
screen "MTA-CFGAvisosBAJA" 1280x800, template "Plantilla"
   TextField "Campo de texto_1" at 477,9 size 354x27; Text 'Configuración de avisos para Baja presión'
   TextField "Campo de texto_9" at 161,54 size 281x34; Text 'Avisos de BAJA PRESIÓN'
   IOField "Campo ES_1" at 295,105 size 130x30; Authorization "Administración de usuarios"; FormatPattern 999.99; Unit  bar
      ProcessValue <- "CFG-BajaHH"
   IOField "Campo ES_2" at 295,240 size 130x31; Authorization "Administración de usuarios"; FormatPattern 9999999; Unit  h
      ProcessValue <- "Varios_HorasMantMC061_1"
   IOField "Campo ES_3" at 295,195 size 130x31; Authorization "Administración de usuarios"; FormatPattern 9999999; Unit  h
      ProcessValue <- "Varios_HorasMantMC060_3"
   IOField "Campo ES_4" at 295,150 size 130x31; Authorization "Administración de usuarios"; FormatPattern 999.99; Unit  bar
      ProcessValue <- "CFG-BajaLL"
   IOField "Campo ES_5" at 295,285 size 130x30; Authorization "Administración de usuarios"; FormatPattern 9999999; Unit  h
      ProcessValue <- "Varios_HorasMantMC061_4"
   IOField "Campo ES_6" at 295,330 size 130x31; Authorization "Administración de usuarios"; FormatPattern 9999999; Unit  h
      ProcessValue <- "Varios_HorasMantMC062_2"
   IOField "Campo ES_7" at 295,375 size 130x31; Authorization "Administración de usuarios"; FormatPattern 9999999; Unit  h
      ProcessValue <- "Varios_HorasMantMC062_5"
   IOField "Campo ES_8" at 295,420 size 130x31; Authorization "Administración de usuarios"; FormatPattern 9999999; Unit  h
      ProcessValue <- "Varios_HorasMantMC063_3"
   TextField "Campo de texto_2" at 15,107 size 293x25; Text 'Presión Aviso límite de presión Máxima'
   TextField "Campo de texto_3" at 15,242 size 238x25; Text 'Tiempo Mant.#1 Comp. Sullair1'
   TextField "Campo de texto_6" at 15,197 size 248x25; Text 'Tiempo Mant. #3 Comp. Sullair2'
   TextField "Campo de texto_4" at 15,152 size 289x25; Text 'Presión Aviso límite de presión Mínima'
   TextField "Campo de texto_5" at 15,287 size 238x25; Text 'Tiempo Mant.#4 Comp. Sullair1'
   TextField "Campo de texto_7" at 15,332 size 238x25; Text 'Tiempo Mant.#2 Comp. Sullair0'
   TextField "Campo de texto_8" at 15,377 size 238x25; Text 'Tiempo Mant.#5 Comp. Sullair0'
   TextField "Campo de texto_10" at 15,422 size 231x25; Text 'Tiempo Mant.#3 Comp. Atlas3'
   IOField "Campo ES_9" at 295,465 size 130x30; Authorization "Administración de usuarios"; FormatPattern 9999999; Unit  h
      ProcessValue <- "Varios_HorasMantMC064_1"
   IOField "Campo ES_10" at 295,510 size 130x31; Authorization "Administración de usuarios"; FormatPattern 9999999; Unit  h
      ProcessValue <- "Varios_HorasMantMC064_4"
   IOField "Campo ES_11" at 295,555 size 130x31; Authorization "Administración de usuarios"; FormatPattern 9999999; Unit  h
      ProcessValue <- "Varios_HorasMantMS054_2"
   TextField "Campo de texto_11" at 15,467 size 231x25; Text 'Tiempo Mant.#1 Comp. Atlas2'
   TextField "Campo de texto_12" at 15,512 size 231x25; Text 'Tiempo Mant.#4 Comp. Atlas2'
   TextField "Campo de texto_13" at 15,557 size 232x25; Text 'Tiempo Mant. #2 Sec. Sullair 1'
   IOField "Campo ES_13" at 716,150 size 130x30; Authorization "Administración de usuarios"; FormatPattern 9999999; Unit  h
      ProcessValue <- "Varios_HorasMantMC060_1"
   IOField "Campo ES_14" at 716,105 size 130x31; Authorization "Administración de usuarios"; FormatPattern 999.99; Unit  bar
      ProcessValue <- "CFG-BajaH"
   IOField "Campo ES_15" at 716,195 size 130x31; Authorization "Administración de usuarios"; FormatPattern 9999999; Unit  h
      ProcessValue <- "Varios_HorasMantMC060_4"
   IOField "Campo ES_16" at 716,240 size 130x31; Authorization "Administración de usuarios"; FormatPattern 9999999; Unit  h
      ProcessValue <- "Varios_HorasMantMC061_2"
   IOField "Campo ES_17" at 716,285 size 130x30; Authorization "Administración de usuarios"; FormatPattern 9999999; Unit  h
      ProcessValue <- "Varios_HorasMantMC061_5"
   IOField "Campo ES_18" at 716,330 size 130x31; Authorization "Administración de usuarios"; FormatPattern 9999999; Unit  h
      ProcessValue <- "Varios_HorasMantMC062_3"
   IOField "Campo ES_19" at 716,375 size 130x31; Authorization "Administración de usuarios"; FormatPattern 9999999; Unit  h
      ProcessValue <- "Varios_HorasMantMC063_1"
   IOField "Campo ES_20" at 716,420 size 130x31; Authorization "Administración de usuarios"; FormatPattern 9999999; Unit  h
      ProcessValue <- "Varios_HorasMantMC063_4"
   TextField "Campo de texto_15" at 436,152 size 248x25; Text 'Tiempo Mant. #1 Comp. Sullair2'
   TextField "Campo de texto_16" at 436,107 size 247x25; Text 'Presión Aviso de presión elevada'
   TextField "Campo de texto_17" at 436,197 size 248x25; Text 'Tiempo Mant. #4 Comp. Sullair2'
   TextField "Campo de texto_18" at 436,242 size 238x25; Text 'Tiempo Mant.#2 Comp. Sullair1'
   TextField "Campo de texto_19" at 436,287 size 238x25; Text 'Tiempo Mant.#5 Comp. Sullair1'
   TextField "Campo de texto_20" at 436,332 size 238x25; Text 'Tiempo Mant.#3 Comp. Sullair0'
   TextField "Campo de texto_21" at 436,377 size 231x25; Text 'Tiempo Mant.#1 Comp. Atlas3'
   TextField "Campo de texto_22" at 436,422 size 231x25; Text 'Tiempo Mant.#4 Comp. Atlas3'
   IOField "Campo ES_21" at 716,465 size 130x30; Authorization "Administración de usuarios"; FormatPattern 9999999; Unit  h
      ProcessValue <- "Varios_HorasMantMC064_2"
   IOField "Campo ES_22" at 716,510 size 130x31; Authorization "Administración de usuarios"; FormatPattern 9999999; Unit  h
      ProcessValue <- "Varios_HorasMantMC064_5"
   IOField "Campo ES_23" at 716,555 size 130x31; Authorization "Administración de usuarios"; FormatPattern 9999999; Unit  h
      ProcessValue <- "Varios_UltimoMantMS055_1"
   TextField "Campo de texto_23" at 436,467 size 231x25; Text 'Tiempo Mant.#2 Comp. Atlas2'
   TextField "Campo de texto_24" at 436,512 size 231x25; Text 'Tiempo Mant.#5 Comp. Atlas2'
   TextField "Campo de texto_25" at 436,557 size 232x25; Text 'Tiempo Mant. #1 Sec. Sullair 2'
   IOField "Campo ES_25" at 1137,195 size 130x30; Authorization "Administración de usuarios"; FormatPattern 9999999; Unit  h
      ProcessValue <- "Varios_UltimoMantMC060_5"
   IOField "Campo ES_26" at 1137,150 size 130x31; Authorization "Administración de usuarios"; FormatPattern 9999999; Unit  h
      ProcessValue <- "Varios_HorasMantMC060_2"
   IOField "Campo ES_27" at 1137,105 size 130x31; Authorization "Administración de usuarios"; FormatPattern 999.99; Unit  bar
      ProcessValue <- "CFG-BajaL"
   IOField "Campo ES_28" at 1137,240 size 130x31; Authorization "Administración de usuarios"; FormatPattern 9999999; Unit  h
      ProcessValue <- "Varios_HorasMantMC061_3"
   IOField "Campo ES_29" at 1137,285 size 130x30; Authorization "Administración de usuarios"; FormatPattern 9999999; Unit  h
      ProcessValue <- "Varios_HorasMantMC062_1"
   IOField "Campo ES_30" at 1137,330 size 130x31; Authorization "Administración de usuarios"; FormatPattern 9999999; Unit  h
      ProcessValue <- "Varios_HorasMantMC062_4"
   IOField "Campo ES_31" at 1137,375 size 130x31; Authorization "Administración de usuarios"; FormatPattern 9999999; Unit  h
      ProcessValue <- "Varios_HorasMantMC063_2"
   IOField "Campo ES_32" at 1137,420 size 130x31; Authorization "Administración de usuarios"; FormatPattern 9999999; Unit  h
      ProcessValue <- "Varios_HorasMantMC063_5"
   TextField "Campo de texto_27" at 857,197 size 243x25; Text 'Tiempo Mant.#5 Comp. Sullair2'
   TextField "Campo de texto_28" at 857,152 size 248x25; Text 'Tiempo Mant. #2 Comp. Sullair2'
   TextField "Campo de texto_29" at 857,107 size 222x25; Text 'Presión Aviso de presión baja'
   TextField "Campo de texto_30" at 857,242 size 238x25; Text 'Tiempo Mant.#3 Comp. Sullair1'
   TextField "Campo de texto_31" at 857,287 size 238x25; Text 'Tiempo Mant.#1 Comp. Sullair0'
   TextField "Campo de texto_32" at 857,332 size 238x25; Text 'Tiempo Mant.#4 Comp. Sullair0'
   TextField "Campo de texto_33" at 857,377 size 231x25; Text 'Tiempo Mant.#2 Comp. Atlas3'
   TextField "Campo de texto_34" at 857,422 size 273x25; Text 'Tiempo mant. #5 compresor Atlas 3'
   IOField "Campo ES_33" at 1137,465 size 130x30; Authorization "Administración de usuarios"; FormatPattern 9999999; Unit  h
      ProcessValue <- "Varios_HorasMantMC064_3"
   IOField "Campo ES_34" at 1137,510 size 130x31; Authorization "Administración de usuarios"; FormatPattern 9999999; Unit  h
      ProcessValue <- "Varios_HorasMantMS054_1"
   IOField "Campo ES_35" at 1137,555 size 130x31; Authorization "Administración de usuarios"; FormatPattern 9999999; Unit  h
      ProcessValue <- "Varios_HorasMantMS055_2"
   TextField "Campo de texto_35" at 857,467 size 231x25; Text 'Tiempo Mant.#3 Comp. Atlas2'
   TextField "Campo de texto_36" at 857,512 size 232x25; Text 'Tiempo Mant. #1 Sec. Sullair 1'
   TextField "Campo de texto_37" at 857,557 size 232x25; Text 'Tiempo Mant. #2 Sec. Sullair 2'

screen "MTA-ChillersBombasEnvasado" 1280x800, template "Plantilla"
   TextField "Campo de texto_5" at 519,10 size 240x27; Text 'Chillers - Bombas Envasado'
   GraphicView "Visor de gráficos_3" at 944,375 size 64x103; Picture "Bomba"
   GraphicIOField "Plantilla_Campo ES gráfico_2" at 980,449 size 81x68; PictureList "Motor2"
      ProcessValue <- "AnimaciónMT009"
   SymbolicIOField "Campo ES simbólico_4" at 890,188 size 220x29; TextOff '0'; TextOn '1'; TextList "EstadoMotor"
      ProcessValue <- "AnimaciónMT009"
   TextField "Campo de texto_6" at 887,129 size 53x23; Text 'MT009'
   GraphicView "Visor de gráficos_4" at 702,375 size 64x103; Picture "Bomba"
   GraphicIOField "Plantilla_Campo ES gráfico_1" at 738,449 size 81x68; PictureList "Motor2"
      ProcessValue <- "AnimaciónMT010"
   SymbolicIOField "Campo ES simbólico_1" at 648,188 size 220x29; TextOff '0'; TextOn '1'; TextList "EstadoMotor"
      ProcessValue <- "AnimaciónMT010"
   TextField "Campo de texto_7" at 645,129 size 53x23; Text 'MT010'
   GraphicView "Visor de gráficos_6" at 216,375 size 64x103; Picture "Bomba"
   GraphicIOField "Plantilla_Campo ES gráfico_4" at 252,449 size 81x68; PictureList "Motor2"
      ProcessValue <- "AnimaciónMP013"
   SymbolicIOField "Campo ES simbólico_3" at 164,188 size 220x29; TextOff '0'; TextOn '1'; TextList "EstadoMotor"
      ProcessValue <- "AnimaciónMP013"
   TextField "Campo de texto_9" at 167,129 size 52x23; Text 'MP013'
   TextField "Campo de texto_19" at 645,160 size 195x18; Text 'Intercambiador Línea 1 y Manomec'
   GraphicView "Visor de gráficos_5" at 460,375 size 64x103; Picture "Bomba"
   GraphicIOField "Plantilla_Campo ES gráfico_3" at 496,449 size 81x68; PictureList "Motor2"
      ProcessValue <- "AnimaciónMP012"
   SymbolicIOField "Campo ES simbólico_2" at 406,188 size 220x29; TextOff '0'; TextOn '1'; TextList "EstadoMotor"
      ProcessValue <- "AnimaciónMP012"
   TextField "Campo de texto_8" at 403,129 size 52x23; Text 'MP012'
   TextField "Campo de texto_18" at 886,160 size 150x18; Text 'Intercambiador Línea 3 y 5'
   TextField "Campo de texto_16" at 407,161 size 150x18; Text 'Chillers Envasado - Principal'
   TextField "Campo de texto_17" at 165,161 size 146x18; Text 'Chillers Envasado - Backup'
   ScreenModuleView "ControlMotor-NoAUTO_1" at 916,230 size 171x108
      Guid_{11997190-67152} <- "DesMT009"
      Guid_{11997190-67156} <- "ParadaMT009"
      Guid_{11997190-67150} <- "HabMT009"
      Guid_{11997190-67154} <- "MarchaMT009"
   ScreenModuleView "ControlMotor-NoAUTO_2" at 676,230 size 171x108
      Guid_{11997190-67152} <- "DesMT010"
      Guid_{11997190-67156} <- "ParadaMT010"
      Guid_{11997190-67150} <- "HabMT010"
      Guid_{11997190-67154} <- "MarchaMT010"
   ScreenModuleView "ControlMotor-NoAUTO_3" at 431,230 size 171x108
      Guid_{11997190-67152} <- "DesMP012"
      Guid_{11997190-67156} <- "ParadaMP012"
      Guid_{11997190-67150} <- "HabMP012"
      Guid_{11997190-67154} <- "MarchaMP012"
   ScreenModuleView "ControlMotor-NoAUTO_4" at 191,230 size 171x108
      Guid_{11997190-67152} <- "DesMP013"
      Guid_{11997190-67156} <- "ParadaMP013"
      Guid_{11997190-67150} <- "HabMP013"
      Guid_{11997190-67154} <- "MarchaMP013"
   Button "Botón_1" at 1184,68 size 48x46; TextOff '?'
      on Click: ActivateScreen("MTA-AyudaMotores", 0)

screen "MTA-ChillersBombasSoplado" 1280x800, template "Plantilla"
   GraphicView "Visor de gráficos_3" at 944,375 size 64x103; Picture "Bomba"
   GraphicView "Visor de gráficos_4" at 702,375 size 64x103; Picture "Bomba"
   GraphicView "Visor de gráficos_6" at 216,375 size 64x103; Picture "Bomba"
   GraphicView "Visor de gráficos_5" at 460,375 size 64x103; Picture "Bomba"
   TextField "Campo de texto_5" at 530,10 size 221x27; Text 'Chillers - Bombas Soplado'
   GraphicIOField "Plantilla_Campo ES gráfico_2" at 980,449 size 81x68; PictureList "Motor2"
      ProcessValue <- "AnimaciónMT007"
   SymbolicIOField "Campo ES simbólico_4" at 890,188 size 220x29; TextOff '0'; TextOn '1'; TextList "EstadoMotor"
      ProcessValue <- "AnimaciónMT007"
   TextField "Campo de texto_6" at 887,129 size 53x23; Text 'MT007'
   GraphicIOField "Plantilla_Campo ES gráfico_1" at 738,449 size 81x68; PictureList "Motor2"
      ProcessValue <- "AnimaciónMT008"
   SymbolicIOField "Campo ES simbólico_1" at 648,188 size 220x29; TextOff '0'; TextOn '1'; TextList "EstadoMotor"
      ProcessValue <- "AnimaciónMT008"
   TextField "Campo de texto_7" at 645,129 size 53x23; Text 'MT008'
   GraphicIOField "Plantilla_Campo ES gráfico_4" at 252,449 size 81x68; PictureList "Motor2"
      ProcessValue <- "AnimaciónMP011"
   SymbolicIOField "Campo ES simbólico_3" at 164,188 size 220x29; TextOff '0'; TextOn '1'; TextList "EstadoMotor"
      ProcessValue <- "AnimaciónMP011"
   TextField "Campo de texto_9" at 167,129 size 52x23; Text 'MP011'
   TextField "Campo de texto_19" at 647,161 size 166x18; Text 'Sopladora Línea 3 y Manomec'
   GraphicIOField "Plantilla_Campo ES gráfico_3" at 496,449 size 81x68; PictureList "Motor2"
      ProcessValue <- "AnimaciónMP010"
   SymbolicIOField "Campo ES simbólico_2" at 406,188 size 220x29; TextOff '0'; TextOn '1'; TextList "EstadoMotor"
      ProcessValue <- "AnimaciónMP010"
   TextField "Campo de texto_8" at 403,129 size 52x23; Text 'MP010'
   TextField "Campo de texto_18" at 887,161 size 104x18; Text 'Sopladora Línea 1'
   TextField "Campo de texto_16" at 404,161 size 142x18; Text 'Chillers Soplado - Principal'
   TextField "Campo de texto_17" at 165,161 size 138x18; Text 'Chillers Soplado - Backup'
   GraphicView "Plantilla_Visor de gráficos_2" at 1232,6 size 35x35; Picture "ParlantesGris_1"
   GraphicView "Plantilla_Visor de gráficos_1" at 1232,6 size 35x35; Picture "ParlantesRojo"
      Visibility <- "SirenaChillers"
   Button "Botón_1" at 1220,1 size 57x44; TextOff 'Text'
      on Click: ActivateScreen("MTA-ChillersCFGSirena", 0)
   ScreenModuleView "ControlMotor-NoAUTO_4" at 916,230 size 171x108
      Guid_{11997190-67152} <- "DesMT007"
      Guid_{11997190-67156} <- "ParadaMT007"
      Guid_{11997190-67150} <- "HabMT007"
      Guid_{11997190-67154} <- "MarchaMT007"
   ScreenModuleView "ControlMotor-NoAUTO_1" at 424,229 size 171x108
      Guid_{11997190-67152} <- "DesMP010"
      Guid_{11997190-67156} <- "ParadaMP010"
      Guid_{11997190-67150} <- "HabMP010"
      Guid_{11997190-67154} <- "MarchaMP010"
   ScreenModuleView "ControlMotor-NoAUTO_2" at 676,230 size 171x108
      Guid_{11997190-67152} <- "DesMT008"
      Guid_{11997190-67156} <- "ParadaMT008"
      Guid_{11997190-67150} <- "HabMT008"
      Guid_{11997190-67154} <- "MarchaMT008"
   ScreenModuleView "ControlMotor-NoAUTO_3" at 184,229 size 171x108
      Guid_{11997190-67152} <- "DesMP011"
      Guid_{11997190-67156} <- "ParadaMP011"
      Guid_{11997190-67150} <- "HabMP011"
      Guid_{11997190-67154} <- "MarchaMP011"
   Button "Botón_2" at 1184,68 size 48x46; TextOff '?'
      on Click: ActivateScreen("MTA-AyudaMotores", 0)

screen "MTA-ChillersCFGSirena" 1280x800, template "Plantilla"
   Switch "Interruptor_1" at 215,155 size 36x32; TextOn 'Habilitado'; TextOff 'Deshabilitado'; CaptionText 'Switch'; PictureOff "ParlantesGrisClaro_1"; Authorization "Administración de usuarios"; PictureOn "ParlantesVerde2_1"
      ProcessValue <- "SirenaM1"
   Switch "Interruptor_2" at 215,192 size 36x32; TextOn 'Habilitado'; TextOff 'Deshabilitado'; CaptionText 'Switch'; PictureOff "ParlantesGrisClaro_1"; Authorization "Administración de usuarios"; PictureOn "ParlantesVerde2_1"
      ProcessValue <- "SirenaM2"
   Switch "Interruptor_3" at 215,229 size 36x32; TextOn 'Habilitado'; TextOff 'Deshabilitado'; CaptionText 'Switch'; PictureOff "ParlantesGrisClaro_1"; Authorization "Administración de usuarios"; PictureOn "ParlantesVerde2_1"
      ProcessValue <- "SirenaM3"
   Switch "Interruptor_4" at 215,266 size 36x32; TextOn 'Habilitado'; TextOff 'Deshabilitado'; CaptionText 'Switch'; PictureOff "ParlantesGrisClaro_1"; Authorization "Administración de usuarios"; PictureOn "ParlantesVerde2_1"
      ProcessValue <- "SirenaM4"
   Switch "Interruptor_5" at 215,303 size 36x32; TextOn 'Habilitado'; TextOff 'Deshabilitado'; CaptionText 'Switch'; PictureOff "ParlantesGrisClaro_1"; Authorization "Administración de usuarios"; PictureOn "ParlantesVerde2_1"
      ProcessValue <- "SirenaM5"
   TextField "Campo de texto_1" at 259,307 size 365x22; Text 'Ninguna Bomba para torres de enfriamiento en marcha'
   TextField "Campo de texto_2" at 259,270 size 424x22; Text 'Ninguna Bomba para Intercambiadores de Envasado en marcha'
   TextField "Campo de texto_3" at 259,234 size 353x22; Text 'Ninguna Bomba para Chillers de Envasado en marcha'
   TextField "Campo de texto_4" at 259,196 size 411x22; Text 'Ninguna Bomba para Intercambiadores de Solpado en marcha'
   TextField "Campo de texto_5" at 259,160 size 340x22; Text 'Ninguna Bomba para Chillers de Soplado en marcha'
   TextField "Campo de texto_6" at 147,93 size 410x22; Text 'Motivos para que la sirena de Chillers se active:'
   Switch "Interruptor_6" at 215,340 size 36x32; TextOn 'Habilitado'; TextOff 'Deshabilitado'; CaptionText 'Switch'; PictureOff "ParlantesGrisClaro_1"; Authorization "Administración de usuarios"; PictureOn "ParlantesVerde2_1"
      ProcessValue <- "SirenaM6"
   TextField "Campo de texto_8" at 259,345 size 231x22; Text 'Ningún Chiller de Soplado Habilitado'
   Switch "Interruptor_7" at 215,377 size 36x32; TextOn 'Habilitado'; TextOff 'Deshabilitado'; CaptionText 'Switch'; PictureOff "ParlantesGrisClaro_1"; Authorization "Administración de usuarios"; PictureOn "ParlantesVerde2_1"
      ProcessValue <- "SirenaM7"
   TextField "Campo de texto_9" at 259,381 size 244x22; Text 'Ningún Chiller de Envasado Habilitado'
   Switch "Interruptor_8" at 215,415 size 36x32; TextOn 'Habilitado'; TextOff 'Deshabilitado'; CaptionText 'Switch'; PictureOff "ParlantesGrisClaro_1"; Authorization "Administración de usuarios"; PictureOn "ParlantesVerde2_1"
      ProcessValue <- "SirenaM8"
   TextField "Campo de texto_10" at 259,420 size 150x22; Text 'Alarma en algún Chiller'
   GraphicView "Plantilla_Visor de gráficos_2" at 1232,6 size 35x35; Picture "ParlantesGris_1"
   GraphicView "Plantilla_Visor de gráficos_1" at 1232,6 size 35x35; Picture "ParlantesRojo"
      Visibility <- "SirenaChillers"
   Button "Botón_1" at 1220,1 size 57x44; TextOff 'Text'
      on Click: ActivateScreen("MTA-ChillersCFGSirena", 0)
   Switch "Interruptor_9" at 215,453 size 36x32; TextOn 'Habilitado'; TextOff 'Deshabilitado'; CaptionText 'Switch'; PictureOff "ParlantesGrisClaro_1"; Authorization "Administración de usuarios"; PictureOn "ParlantesVerde2_1"
      ProcessValue <- "SirenaM9"
   TextField "Campo de texto_11" at 259,458 size 194x22; Text 'Falla Térmica en algún motor'
   TextField "Campo de texto_7" at 505,9 size 270x27; Text 'Configuración de Sirena Chillers'

screen "MTA-Chillers-General" 1280x800, template "Plantilla"
   GraphicView "Visor de gráficos_7" at 774,285 size 48x87; Picture "Bomba"
   GraphicView "Visor de gráficos_8" at 838,285 size 48x87; Picture "Bomba"
   GraphicView "Visor de gráficos_1" at 646,285 size 48x87; Picture "Bomba"
   GraphicView "Visor de gráficos_9" at 710,285 size 48x87; Picture "Bomba"
   GraphicView "Visor de gráficos_3" at 1155,429 size 120x284; Picture "Chiller2bb"
   GraphicView "Visor de gráficos_4" at 950,233 size 168x168; Picture "Chiller_2"
   GraphicView "Visor de gráficos_5" at 494,285 size 48x87; Picture "Bomba"
   GraphicView "Visor de gráficos_6" at 558,285 size 48x87; Picture "Bomba"
   GraphicView "Visor de gráficos_10" at 366,285 size 48x87; Picture "Bomba"
   GraphicView "Visor de gráficos_11" at 430,285 size 48x87; Picture "Bomba"
   GraphicView "Visor de gráficos_2" at 12,188 size 200x216; Picture "Chiller2b"
   GraphicView "Visor de gráficos_12" at 107,550 size 160x149; Picture "Chillerb"
   GraphicView "Visor de gráficos_15" at 351,213 size 116x103; Picture "tubo"
   GraphicView "Visor de gráficos_16" at 479,213 size 116x103; Picture "tubo"
   GraphicView "Visor de gráficos_17" at 631,213 size 116x103; Picture "tubo"
   GraphicView "Visor de gráficos_18" at 759,213 size 116x103; Picture "tubo"
   GraphicView "Visor de gráficos_14" at 622,54 size 245x227; Picture "Tanque3_1"
   GraphicView "Visor de gráficos_13" at 344,46 size 245x227; Picture "Tanque3_1"
   GraphicView "Plantilla_Visor de gráficos_2" at 1232,6 size 35x35; Picture "ParlantesGris_1"
   GraphicView "Plantilla_Visor de gráficos_1" at 1232,6 size 35x35; Picture "ParlantesRojo"
      Visibility <- "SirenaChillers"
   GraphicIOField "Plantilla_Campo ES gráfico_2" at 529,355 size 57x52; PictureList "Motor2"
      ProcessValue <- "AnimaciónMT010"
   GraphicIOField "Plantilla_Campo ES gráfico_1" at 593,355 size 57x52; PictureList "Motor2"
      ProcessValue <- "AnimaciónMT009"
   GraphicIOField "Plantilla_Campo ES gráfico_3" at 809,355 size 57x52; PictureList "Motor2"
      ProcessValue <- "AnimaciónMT008"
   GraphicIOField "Plantilla_Campo ES gráfico_4" at 873,355 size 57x52; PictureList "Motor2"
      ProcessValue <- "AnimaciónMT007"
   GraphicIOField "Plantilla_Campo ES gráfico_5" at 681,355 size 57x52; PictureList "Motor2"
      ProcessValue <- "AnimaciónMP011"
   GraphicIOField "Plantilla_Campo ES gráfico_6" at 745,355 size 57x52; PictureList "Motor2"
      ProcessValue <- "AnimaciónMP010"
   GraphicIOField "Plantilla_Campo ES gráfico_7" at 401,355 size 57x52; PictureList "Motor2"
      ProcessValue <- "AnimaciónMP013"
   GraphicIOField "Plantilla_Campo ES gráfico_8" at 465,355 size 57x52; PictureList "Motor2"
      ProcessValue <- "AnimaciónMP012"
   TextField "Campo de texto_1" at 984,196 size 86x32; Text 'Chiller Soplado Chico'
   TextField "Campo de texto_2" at 1027,485 size 86x32; Text 'Chiller Soplado Grande'
   TextField "Campo de texto_3" at 134,514 size 90x32; Text 'Chiller Envasado Chico'
   TextField "Campo de texto_4" at 60,150 size 90x32; Text 'Chiller Envasado Grande'
   TextField "Campo de texto_6" at 762,451 size 131x25; Text 'Bombas Soplado'
   TextField "Campo de texto_7" at 477,451 size 139x25; Text 'Bombas Envasado'
   TextField "Campo de texto_9" at 848,132 size 51x52; Text 'Tanque Soplado'
   TextField "Campo de texto_8" at 424,419 size 41x19; Text 'MP013'
   TextField "Campo de texto_11" at 485,419 size 41x19; Text 'MP012'
   TextField "Campo de texto_12" at 546,419 size 49x19; Text 'MT010'
   TextField "Campo de texto_13" at 614,419 size 42x19; Text 'MT009'
   TextField "Campo de texto_14" at 703,419 size 41x19; Text 'MP011'
   TextField "Campo de texto_15" at 767,419 size 41x19; Text 'MP010'
   TextField "Campo de texto_16" at 830,419 size 42x19; Text 'MT008'
   TextField "Campo de texto_17" at 893,419 size 42x19; Text 'MT007'
   TextField "Campo de texto_10" at 569,131 size 58x52; Text 'Tanque Envasado'
   TextField "Campo de texto_21" at 242,362 size 40x18; Text 'Alarma'
   TextField "Campo de texto_22" at 242,341 size 108x18; Text 'En Funcionamiento'
   TextField "Campo de texto_23" at 242,382 size 101x18; Text 'Máxima Capacidad'
   TextField "Campo de texto_24" at 299,638 size 79x18; Text 'Alarma Aceite'
   TextField "Campo de texto_25" at 299,617 size 108x18; Text 'En Funcionamiento'
   TextField "Campo de texto_26" at 299,660 size 115x18; Text 'Alarma Temperatura'
   TextField "Campo de texto_27" at 299,681 size 125x18; Text 'Alarma Térmico motor'
   TextField "Campo de texto_18" at 1037,602 size 40x18; Text 'Alarma'
   TextField "Campo de texto_19" at 1037,581 size 108x18; Text 'En Funcionamiento'
   TextField "Campo de texto_20" at 1037,622 size 101x18; Text 'Máxima Capacidad'
   TextField "Campo de texto_28" at 1154,313 size 120x18; Text 'Motor 2 Funcionando'
   TextField "Campo de texto_29" at 1154,292 size 120x18; Text 'Motor 1 Funcionando'
   TextField "Campo de texto_30" at 1154,335 size 96x18; Text 'Térmico motor 1'
   TextField "Campo de texto_31" at 1154,356 size 96x18; Text 'Térmico motor 2'
   Button "Botón_2" at 657,329 size 295x86; TextOff 'Control Soplado'
      on Click: ActivateScreen("MTA-ChillersBombasSoplado", 0)
   Button "Botón_5" at 361,328 size 296x87; TextOff 'Control Envasado'
      on Click: ActivateScreen("MTA-ChillersBombasEnvasado", 0)
   Button "Botón_1" at 1220,1 size 57x44; TextOff 'Text'
      on Click: ActivateScreen("MTA-ChillersCFGSirena", 0)
   Switch "Interruptor_1" at 222,294 size 91x31; TextOn 'Deshabilitado'; TextOff 'Habilitado'; CaptionText 'Switch'; Authorization "Administración de usuarios"
      Appearance <- "Habilitación-CH-ENV-GR"
      ProcessValue <- "Habilitación-CH-ENV-GR"
   Switch "Interruptor_2" at 279,570 size 91x31; TextOn 'Deshabilitado'; TextOff 'Habilitado'; CaptionText 'Switch'; Authorization "Administración de usuarios"
      Appearance <- "Habilitación-CH-ENV-CH"
      ProcessValue <- "Habilitación-CH-ENV-CH"
   Switch "Interruptor_3" at 1017,534 size 91x31; TextOn 'Deshabilitado'; TextOff 'Habilitado'; CaptionText 'Switch'; Authorization "Administración de usuarios"
      Appearance <- "Habilitación-CH-SOP-GR"
      ProcessValue <- "Habilitación-CH-SOP-GR"
   Switch "Interruptor_4" at 1135,252 size 91x31; TextOn 'Deshabilitado'; TextOff 'Habilitado'; CaptionText 'Switch'; Authorization "Administración de usuarios"
      Appearance <- "Habilitación-CH-SOP-CH"
      ProcessValue <- "Habilitación-CH-SOP-CH"
   Circle "Círculo_1" at 222,384 size 16x16
      Appearance <- "MAX-CH-ENV-GR"
   Circle "Círculo_10" at 222,342 size 16x16
      Appearance <- "RUN-CH-ENV-GR"
   Circle "Círculo_11" at 222,363 size 16x16
      Appearance <- "Alarma1-CH-ENV-GR"
   Circle "Círculo_2" at 279,618 size 16x16
      Appearance <- "CH-ENV-CH-RUN"
   Circle "Círculo_3" at 279,639 size 16x16
      Appearance <- "CH-ENV-CH-ACT"
   Circle "Círculo_5" at 279,661 size 16x16
      Appearance <- "CH-ENV-CH-TEMP"
   Circle "Círculo_6" at 279,682 size 16x16
      Appearance <- "CH-ENV-CH-TERM"
   Circle "Círculo_4" at 1016,624 size 16x16
      Appearance <- "MAX-CH-SOP-GR"
   Circle "Círculo_7" at 1016,581 size 16x16
      Appearance <- "RUN-CH-SOP-GR"
   Circle "Círculo_8" at 1016,603 size 16x16
      Appearance <- "Alarma1-CH-SOP-GR"
   Circle "Círculo_9" at 1132,293 size 16x16
      Appearance <- "CH-SOP-CH-CTC1ON"
   Circle "Círculo_12" at 1132,314 size 16x16
      Appearance <- "CH-SOP-CH-CTC2ON"
   Circle "Círculo_13" at 1132,336 size 16x16
      Appearance <- "CH-SOP-CH-TERM1"
   Circle "Círculo_14" at 1132,357 size 16x16
      Appearance <- "CH-SOP-CH-TERM2"
   Button "Botón_3" at 1184,68 size 48x46; TextOff '?'
      on Click: ActivateScreen("MTA-AyudaColores", 0)
   TextField "Campo de texto_32" at 610,9 size 63x27; Text 'Chillers'

screen "MTA-CompBAJA" 1280x800, template "Plantilla"
   GraphicIOField "Campo ES gráfico_10" at 491,153 size 189x58; PictureList "BaseSullChico"
      ProcessValue <- "AnimaMC064"
   GraphicIOField "Campo ES gráfico_9" at 427,241 size 189x58; PictureList "BaseSullChico"
      ProcessValue <- "AnimaMC063"
   GraphicIOField "Campo ES gráfico_7" at 387,316 size 178x52; PictureList "BaseSullChico"
      ProcessValue <- "AnimaMC062"
   GraphicIOField "Campo ES gráfico_6" at 340,387 size 178x52; PictureList "BaseSullChico"
      ProcessValue <- "AnimaMC061"
   GraphicIOField "Campo ES gráfico_8" at 275,454 size 197x58; PictureList "BaseSullChico"
      ProcessValue <- "AnimaMC060"
   GraphicView "Visor de gráficos_1" at 467,72 size 269x127; Picture "Baja1X_1"
   GraphicView "Visor de gráficos_7" at 467,72 size 269x127; Picture "Baja1Xd"
      Visibility <- "MantM064"
   GraphicView "Visor de gráficos_2" at 403,160 size 269x127; Picture "Baja1X_1"
   GraphicView "Visor de gráficos_8" at 403,160 size 269x127; Picture "Baja1Xd"
      Visibility <- "MantM063"
   GraphicView "Visor de gráficos_3" at 315,232 size 269x127; Picture "baja2X_2"
   GraphicView "Visor de gráficos_9" at 315,232 size 269x127; Picture "baja2Xd_1"
      Visibility <- "MantM062"
   GraphicView "Visor de gráficos_4" at 267,304 size 269x127; Picture "baja2X_2"
   GraphicView "Visor de gráficos_10" at 267,304 size 269x127; Picture "baja2Xd_1"
      Visibility <- "MantM061"
   GraphicView "Visor de gráficos_5" at 243,376 size 213x127; Picture "baja3X_2"
   GraphicView "Visor de gráficos_11" at 243,376 size 213x127; Picture "baja3Xd"
      Visibility <- "MantM060"
   GraphicView "Visor de gráficos_6" at 132,415 size 202x177; Picture "tanque2X_2"
   IOField "Campo ES_1" at 161,449 size 148x28; FormatPattern s999.9; Unit  bar
      ProcessValue <- "PresiónBAJA"
   Button "Botón_3" at 1184,48 size 48x46; TextOff '?'
      on Click: ActivateScreen("MTA-AyudaCmpBaja", 0)
   Button "Botón_1" at 35,197 size 160x46; TextOff 'CFG Avisos'
      on Click: ActivateScreen("MTA-CFGAvisosBAJA", 0)
   TextField "Campo de texto_1" at 516,9 size 248x27; Text 'Compresores de Baja presión'
   GraphicView "Visor de gráficos_12" at 18,528 size 229x141; Picture "Booster-A"
   GraphicIOField "Campo ES gráfico_11" at 68,583 size 48x46; PictureList "Motor Grande"
      ProcessValue <- "AnimaMotBooster"
   GraphicIOField "Campo ES gráfico_12" at 160,500 size 17x32; PictureList "Motor Chico"
      ProcessValue <- "AnimaMotBooster"
   GraphicIOField "Campo ES gráfico_13" at 40,563 size 169x87; PictureList "Hélice"
      ProcessValue <- "Booster_Conf_Marcha"
   GraphicView "Visor de gráficos_18" at 440,520 size 40x40; Picture "MECH2"
   GraphicView "Visor de gráficos_19" at 440,520 size 40x40; Picture "MECH1"
      Visibility <- "Booster2_ModoManten"
   Button "Botón_11" at 440,520 size 40x40; TextOff 'Text'; PictureList "Mantenimiento"
      on Release: SetBit("Booster2_PlsManten")
   GraphicView "Visor de gráficos_17" at 226,528 size 229x141; Picture "Booster-A"
   GraphicIOField "Campo ES gráfico_15" at 286,586 size 48x47; PictureList "Motor Grande"
      ProcessValue <- "AnimaMotBooster2"
   GraphicIOField "Campo ES gráfico_16" at 368,500 size 18x34; PictureList "Motor Chico"
      ProcessValue <- "AnimaMotBooster2"
   GraphicIOField "Campo ES gráfico_17" at 261,565 size 156x84; PictureList "Hélice"
      ProcessValue <- "Booster2_Conf_Marcha"
   GraphicView "Visor de gráficos_13" at 37,520 size 40x40; Picture "MECH2"
   GraphicView "Visor de gráficos_14" at 37,520 size 40x40; Picture "MECH1"
      Visibility <- "Booster_ModoManten"
   Button "Botón_6" at 37,520 size 40x40; TextOff 'Text'; PictureList "Mantenimiento"
      on Release: SetBit("Booster_PlsManten")
   TextField "Campo de texto_4" at 48,674 size 122x19; Text 'Prioridad Marcha'
      Visibility <- "PrioridadBoost1"
   TextField "Campo de texto_10" at 251,674 size 122x19; Text 'Prioridad Marcha'
      Visibility <- "PrioridadBoost2"
   GraphicIOField "Campo ES gráfico_1" at 712,259 size 507x6; PictureList "Indicador"
      ProcessValue <- "AnimaMC063"
   GraphicIOField "Campo ES gráfico_2" at 665,347 size 507x6; PictureList "Indicador"
      ProcessValue <- "AnimaMC062"
   GraphicIOField "Campo ES gráfico_3" at 616,435 size 510x6; PictureList "Indicador"
      ProcessValue <- "AnimaMC061"
   GraphicIOField "Campo ES gráfico_4" at 568,524 size 511x6; PictureList "Indicador"
      ProcessValue <- "AnimaMC060"
   GraphicIOField "Campo ES gráfico_5" at 761,172 size 507x6; PictureList "Indicador"
      ProcessValue <- "AnimaMC064"
   TextField "Campo de texto_5" at 593,449 size 116x39; Text 'Sullair 2'
   TextField "Campo de texto_6" at 641,361 size 116x39; Text 'Sullair 1'
   TextField "Campo de texto_7" at 689,273 size 116x39; Text 'Sullair 0'
   TextField "Campo de texto_8" at 729,185 size 91x39; Text 'Atlas 3'
   TextField "Campo de texto_9" at 785,97 size 100x39; Text 'Atlas 2'
   SymbolicIOField "Campo ES simbólico_5" at 787,133 size 242x21; TextOff '0'; TextOn '1'; TextList "EstadoMotor"
      ProcessValue <- "AnimaMC064"
   SymbolicIOField "Campo ES simbólico_6" at 731,221 size 242x21; TextOff '0'; TextOn '1'; TextList "EstadoMotor"
      ProcessValue <- "AnimaMC063"
   SymbolicIOField "Campo ES simbólico_7" at 691,309 size 242x21; TextOff '0'; TextOn '1'; TextList "EstadoMotor"
      ProcessValue <- "AnimaMC062"
   SymbolicIOField "Campo ES simbólico_8" at 643,397 size 242x21; TextOff '0'; TextOn '1'; TextList "EstadoMotor"
      ProcessValue <- "AnimaMC061"
   SymbolicIOField "Campo ES simbólico_9" at 595,485 size 242x21; TextOff '0'; TextOn '1'; TextList "EstadoMotor"
      ProcessValue <- "AnimaMC060"
   IOField "Campo ES_6" at 595,505 size 85x19; FormatPattern 999999999; Unit  hs
      ProcessValue <- "HorasCmpBaja_HMMC060"
      Appearance <- "EstadoMantMC060"
   IOField "Campo ES_4" at 643,416 size 85x19; FormatPattern 999999999; Unit  hs
      Appearance <- "EstadoMantMC061"
      ProcessValue <- "HorasCmpBaja_HMMC061"
   IOField "Campo ES_5" at 691,328 size 85x19; FormatPattern 999999999; Unit  hs
      ProcessValue <- "HorasCmpBaja_HMMC062"
      Appearance <- "EstadoMantMC062"
   IOField "Campo ES_7" at 731,240 size 85x19; FormatPattern 999999999; Unit  hs
      ProcessValue <- "HorasCmpBaja_HMMC063"
      Appearance <- "EstadoMantMC063"
   IOField "Campo ES_8" at 787,152 size 85x19; FormatPattern 999999999; Unit  hs
      Appearance <- "EstadoMantMC064"
      ProcessValue <- "HorasCmpBaja_HMMC064"
   Switch "Interruptor_1" at 983,102 size 29x29; TextOn '1'; TextOff '0'; CaptionText 'Switch'; PictureOff "A2"; Authorization "Operación"; PictureOn "A"
      ProcessValue <- "AutoMC064"
      Visibility <- "MantM064"
   Switch "Interruptor_2" at 933,190 size 29x29; TextOn '1'; TextOff '0'; CaptionText 'Switch'; PictureOff "A2"; Authorization "Operación"; PictureOn "A"
      ProcessValue <- "AutoMC063"
      Visibility <- "MantM063"
   Switch "Interruptor_3" at 888,278 size 29x29; TextOn '1'; TextOff '0'; CaptionText 'Switch'; PictureOff "A2"; Authorization "Operación"; PictureOn "A"
      ProcessValue <- "AutoMC062"
      Visibility <- "MantM062"
   Switch "Interruptor_4" at 844,367 size 29x29; TextOn '1'; TextOff '0'; CaptionText 'Switch'; PictureOff "A2"; Authorization "Operación"; PictureOn "A"
      ProcessValue <- "AutoMC061"
      Visibility <- "MantM061"
   ScreenModuleView "Faceplate_1_1" at 888,370 size 236x58
      Guid_{11997190-23979} <- "HabilitaciónMC061"
      Guid_{11997190-23983} <- "ParadaMC061"
      Guid_{11997190-23981} <- "MarchaMC061"
      Guid_{11997190-23989} <- "SpoffMC061"
      Guid_{11997190-23976} <- "DeshabilitaciónMC061"
      Guid_{11997190-23987} <- "SponMC061"
      Guid_{11997190-23985} <- "AnimMenuMC061"
   ScreenModuleView "Faceplate_1_3" at 931,281 size 236x58
      Guid_{11997190-23979} <- "HabilitaciónMC062"
      Guid_{11997190-23983} <- "ParadaMC062"
      Guid_{11997190-23981} <- "MarchaMC062"
      Guid_{11997190-23989} <- "SpoffMC062"
      Guid_{11997190-23976} <- "DeshabilitaciónMC062"
      Guid_{11997190-23987} <- "SponMC062"
      Guid_{11997190-23985} <- "AnimMenuMC062"
   ScreenModuleView "Faceplate_1_4" at 980,192 size 236x58
      Guid_{11997190-23979} <- "HabilitaciónMC063"
      Guid_{11997190-23983} <- "ParadaMC063"
      Guid_{11997190-23981} <- "MarchaMC063"
      Guid_{11997190-23989} <- "SpoffMC063"
      Guid_{11997190-23976} <- "DeshabilitaciónMC063"
      Guid_{11997190-23987} <- "SponMC063"
      Guid_{11997190-23985} <- "AnimMenuMC063"
   ScreenModuleView "Faceplate_1_5" at 1030,105 size 236x58
      Guid_{11997190-23979} <- "HabilitaciónMC064"
      Guid_{11997190-23983} <- "ParadaMC064"
      Guid_{11997190-23981} <- "MarchaMC064"
      Guid_{11997190-23989} <- "SpoffMC064"
      Guid_{11997190-23976} <- "DeshabilitaciónMC064"
      Guid_{11997190-23987} <- "SponMC064"
      Guid_{11997190-23985} <- "AnimMenuMC064"
   Switch "Interruptor_6" at 313,243 size 40x40; TextOn '1'; TextOff '0'; CaptionText 'Switch'; PictureOff "MECH2"; PictureOn "MECH1"
      ProcessValue <- "MantM062"
   Switch "Interruptor_7" at 265,323 size 40x40; TextOn '1'; TextOff '0'; CaptionText 'Switch'; PictureOff "MECH2"; PictureOn "MECH1"
      ProcessValue <- "MantM061"
   Switch "Interruptor_9" at 365,171 size 40x40; TextOn '1'; TextOff '0'; CaptionText 'Switch'; PictureOff "MECH2"; PictureOn "MECH1"
      ProcessValue <- "MantM063"
   Switch "Interruptor_10" at 429,83 size 40x40; TextOn '1'; TextOff '0'; CaptionText 'Switch'; PictureOff "MECH2"; PictureOn "MECH1"
      ProcessValue <- "MantM064"
   Switch "Interruptor_5" at 930,472 size 91x31; TextOn 'Deshabilitado'; TextOff 'Habilitado'; CaptionText 'Switch'; Authorization "Administración de usuarios"
      Appearance <- "HabilitarMC060"
      ProcessValue <- "HabilitarMC060"
   Button "Botón_14" at 568,449 size 262x74; TextOff 'Text'
      on Click: ActivateScreen("EPROC-BAJAMC060", 0)
   Button "Botón_15" at 616,361 size 200x74; TextOff 'Text'
      on Click: ActivateScreen("EPROC-BAJAMC061", 0)
   Button "Botón_16" at 664,273 size 200x74; TextOff 'Text'
      on Click: ActivateScreen("EPROC-BAJAMC062", 0)
   Button "Botón_17" at 712,185 size 200x74; TextOff 'Text'
      on Click: ActivateScreen("EPROC-BAJAMC063", 0)
   Button "Botón_18" at 760,97 size 200x74; TextOff 'Text'
      on Click: ActivateScreen("EPROC-BAJAMC064", 0)

screen "MTA-SecALTA" 1280x800, template "Plantilla"
   GraphicIOField "Campo ES gráfico_4" at 981,258 size 280x222; PictureList "Secador1"
      ProcessValue <- "AnimaMS050"
   GraphicView "Visor de gráficos_4" at 999,137 size 234x314; Picture "secador4"
   GraphicView "Visor de gráficos_15" at 999,137 size 234x314; Picture "secador4d_1"
      Visibility <- "MantMS050"
   GraphicIOField "Campo ES gráfico_8" at 571,212 size 366x99; PictureList "Secador2"
      ProcessValue <- "AnimaMS053"
   GraphicView "Visor de gráficos_3" at 592,100 size 363x184; Picture "secador2_3"
   GraphicView "Visor de gráficos_5" at 592,100 size 363x184; Picture "secador2m_1"
      Visibility <- "MantMS053"
   GraphicIOField "Campo ES gráfico_7" at 674,357 size 309x81; PictureList "Secador2"
      ProcessValue <- "AnimaMS052"
   GraphicView "Visor de gráficos_2" at 696,255 size 292x158; Picture "secador3_1"
   GraphicView "Visor de gráficos_6" at 695,255 size 294x158; Picture "secador3d_1"
      Visibility <- "MantMS052"
   GraphicIOField "Campo ES gráfico_6" at 765,490 size 338x86; PictureList "Secador2"
      ProcessValue <- "AnimaMS051"
   GraphicView "Visor de gráficos_1" at 786,405 size 292x142; Picture "secador3_3"
   GraphicView "Visor de gráficos_14" at 786,405 size 292x142; Picture "secador3d_2"
      Visibility <- "MantMS051"
   Button "Botón_3" at 1184,68 size 48x46; TextOff '?'
      on Click: ActivateScreen("MTA-AyudaSecAlta", 0)
   TextField "Campo de texto_7" at 530,9 size 221x27; Text 'Secadores de Alta presión'
   GraphicIOField "Campo ES gráfico_9" at 197,577 size 511x6; PictureList "Indicador"
      ProcessValue <- "AnimaMS051"
   TextField "Campo de texto_6" at 222,499 size 89x39; Text 'ABC 3'
   SymbolicIOField "Campo ES simbólico_9" at 224,535 size 242x21; TextOff '0'; TextOn '1'; TextList "EstadoMotor"
      ProcessValue <- "AnimaMS051"
   GraphicIOField "Campo ES gráfico_1" at 101,439 size 511x6; PictureList "Indicador"
      ProcessValue <- "AnimaMS052"
   TextField "Campo de texto_1" at 126,361 size 89x39; Text 'ABC 2'
   SymbolicIOField "Campo ES simbólico_1" at 128,397 size 242x21; TextOff '0'; TextOn '1'; TextList "EstadoMotor"
      ProcessValue <- "AnimaMS052"
   GraphicIOField "Campo ES gráfico_2" at 21,303 size 511x6; PictureList "Indicador"
      ProcessValue <- "AnimaMS053"
   TextField "Campo de texto_2" at 46,220 size 101x39; Text 'Fargon'
   SymbolicIOField "Campo ES simbólico_2" at 48,256 size 242x21; TextOff '0'; TextOn '1'; TextList "EstadoMotor"
      ProcessValue <- "AnimaMS053"
   GraphicIOField "Campo ES gráfico_3" at 741,681 size 511x6; PictureList "Indicador"
      ProcessValue <- "AnimaMS050"
   TextField "Campo de texto_3" at 766,603 size 89x39; Text 'ABC 1'
   SymbolicIOField "Campo ES simbólico_3" at 768,639 size 242x21; TextOff '0'; TextOn '1'; TextList "EstadoMotor"
      ProcessValue <- "AnimaMS050"
   IOField "Campo ES_6" at 51,282 size 85x19; FormatPattern 999999999; Unit  hs
      ProcessValue <- "HorasSecAlta_HMMS053"
      Appearance <- "LimiteMantMS053"
   IOField "Campo ES_1" at 131,418 size 85x19; FormatPattern 999999999; Unit  hs
      ProcessValue <- "HorasSecAlta_HMMS052"
      Appearance <- "LimiteMantMS052"
   IOField "Campo ES_2" at 227,558 size 85x19; FormatPattern 999999999; Unit  hs
      ProcessValue <- "HorasSecAlta_HMMS051"
      Appearance <- "LimiteMantMS051"
   IOField "Campo ES_3" at 771,660 size 85x19; FormatPattern 999999999; Unit  hs
      ProcessValue <- "HorasSecAlta_HMMS050"
      Appearance <- "LimiteMantMS050"
   Switch "Interruptor_1" at 640,315 size 40x40; TextOn '1'; TextOff '0'; CaptionText 'Switch'; PictureOff "MECH2"; PictureOn "MECH1"
      ProcessValue <- "MantMS052"
   Switch "Interruptor_2" at 731,440 size 40x40; TextOn '1'; TextOff '0'; CaptionText 'Switch'; PictureOff "MECH2"; PictureOn "MECH1"
      ProcessValue <- "MantMS051"
   Switch "Interruptor_3" at 540,176 size 40x40; TextOn '1'; TextOff '0'; CaptionText 'Switch'; PictureOff "MECH2"; PictureOn "MECH1"
      ProcessValue <- "MantMS053"
   Switch "Interruptor_4" at 1212,488 size 40x40; TextOn '1'; TextOff '0'; CaptionText 'Switch'; PictureOff "MECH2"; PictureOn "MECH1"
      ProcessValue <- "MantMS050"
   Switch "Interruptor_5" at 387,506 size 29x29; TextOn '1'; TextOff '0'; CaptionText 'Switch'; PictureOff "A2"; Authorization "Operación"; PictureOn "A"
      ProcessValue <- "AutoMS051"
      Visibility <- "MantMS051"
   Switch "Interruptor_6" at 307,370 size 29x29; TextOn '1'; TextOff '0'; CaptionText 'Switch'; PictureOff "A2"; Authorization "Operación"; PictureOn "A"
      ProcessValue <- "AutoMS052"
      Visibility <- "MantMS052"
   Switch "Interruptor_7" at 227,229 size 29x29; TextOn '1'; TextOff '0'; CaptionText 'Switch'; PictureOff "A2"; Authorization "Operación"; PictureOn "A"
      ProcessValue <- "AutoMS053"
      Visibility <- "MantMS053"
   Switch "Interruptor_8" at 925,606 size 29x29; TextOn '1'; TextOff '0'; CaptionText 'Switch'; PictureOff "A2"; Authorization "Operación"; PictureOn "A"
      ProcessValue <- "AutoMS050"
      Visibility <- "MantMS050"
   ScreenModuleView "Faceplate_2_1" at 453,489 size 244x69
      Guid_{11997190-23979} <- "HabilitaciónMS051"
      Guid_{11997190-37146} <- "Enc1MS051"
      Guid_{11997190-23983} <- "ParadaMS051"
      Guid_{11997190-23981} <- "MarchaMS051"
      Guid_{11997190-37150} <- "Enc2MS051"
      Guid_{11997190-23976} <- "DeshabilitaciónMS051"
      Guid_{11997190-23985} <- "AnimaMenuMS051"
   ScreenModuleView "Faceplate_2_2" at 357,351 size 244x69
      Guid_{11997190-23979} <- "HabilitaciónMS052"
      Guid_{11997190-37146} <- "Enc1MS052"
      Guid_{11997190-23983} <- "ParadaMS052"
      Guid_{11997190-23981} <- "MarchaMS052"
      Guid_{11997190-37150} <- "Enc2MS052"
      Guid_{11997190-23976} <- "DeshabilitaciónMS052"
      Guid_{11997190-23985} <- "AnimaMenuMS052"
   ScreenModuleView "Faceplate_2_3" at 276,215 size 244x69
      Guid_{11997190-23979} <- "HabilitaciónMS053"
      Guid_{11997190-37146} <- "Enc1MS053"
      Guid_{11997190-23983} <- "ParadaMS053"
      Guid_{11997190-23981} <- "MarchaMS053"
      Guid_{11997190-37150} <- "Enc2MS053"
      Guid_{11997190-23976} <- "DeshabilitaciónMS053"
      Guid_{11997190-23985} <- "AnimaMenuMS053"
   ScreenModuleView "Faceplate_2_4" at 994,593 size 244x69
      Guid_{11997190-23979} <- "HabilitaciónMS050"
      Guid_{11997190-37146} <- "Enc1MS050"
      Guid_{11997190-23983} <- "ParadaMS050"
      Guid_{11997190-23981} <- "MarchaMS050"
      Guid_{11997190-37150} <- "Enc2MS050"
      Guid_{11997190-23976} <- "DeshabilitaciónMS050"
      Guid_{11997190-23985} <- "AnimaMenuMS050"
   Button "Botón_1" at 741,590 size 150x90; TextOff 'Text'
      on Click: ActivateScreen("EPROC-ALTAMS050", 0)
   Button "Botón_2" at 197,486 size 150x90; TextOff 'Text'
      on Click: ActivateScreen("EPROC-ALTAMS051", 0)
   Button "Botón_4" at 101,348 size 150x90; TextOff 'Text'
      on Click: ActivateScreen("EPROC-ALTAMS052", 0)
   Button "Botón_5" at 21,212 size 150x90; TextOff 'Text'
      on Click: ActivateScreen("EPROC-ALTAMS053", 0)

screen "MTA-SecBaja" 1280x800, template "Plantilla"
   GraphicIOField "Campo ES gráfico_4" at 639,360 size 511x6; PictureList "Indicador"
      ProcessValue <- "AnimaMS055"
   TextField "Campo de texto_5" at 664,282 size 116x39; Text 'Sullair 2'
   SymbolicIOField "Campo ES simbólico_9" at 666,318 size 242x21; TextOff '0'; TextOn '1'; TextList "EstadoMotor"
      ProcessValue <- "AnimaMS055"
   GraphicIOField "Campo ES gráfico_3" at 482,493 size 510x6; PictureList "Indicador"
      ProcessValue <- "AnimaMS054"
   TextField "Campo de texto_6" at 507,415 size 116x39; Text 'Sullair 1'
   SymbolicIOField "Campo ES simbólico_8" at 509,451 size 242x21; TextOff '0'; TextOn '1'; TextList "EstadoMotor"
      ProcessValue <- "AnimaMS054"
   IOField "Campo ES_6" at 666,339 size 85x19; FormatPattern 999999999; Unit  hs
      Appearance <- "EstadoMantMC060"
      ProcessValue <- "HorasSecBaja_HMMS055"
   IOField "Campo ES_1" at 509,472 size 85x19; FormatPattern 999999999; Unit  hs
      Appearance <- "EstadoMantMC060"
      ProcessValue <- "HorasSecBaja_HMMS054"
   ScreenModuleView "Faceplate_3_2" at 923,282 size 213x73; ScreenModuleType ""
      Guid_{11997190-23981} <- "MarchaMS055"
      Guid_{11997190-23979} <- "HabilitaciónMS055"
      Guid_{11997190-23976} <- "DeshabilitaciónMS055"
      Guid_{11997190-23983} <- "ParadaMS055"
   ScreenModuleView "Faceplate_3_1" at 761,415 size 213x73; ScreenModuleType ""
      Guid_{11997190-23981} <- "MarchaMS054"
      Guid_{11997190-23979} <- "HabilitaciónMS054"
      Guid_{11997190-23976} <- "DeshabilitaciónMS054"
      Guid_{11997190-23983} <- "ParadaMS054"
   Switch "Interruptor_7" at 271,262 size 40x40; TextOn '1'; TextOff '0'; CaptionText 'Switch'; PictureOff "MECH2"; Authorization "Operación"; PictureOn "MECH1"
      ProcessValue <- "MantMS055"
   Switch "Interruptor_8" at 131,406 size 40x40; TextOn '1'; TextOff '0'; CaptionText 'Switch'; PictureOff "MECH2"; Authorization "Operación"; PictureOn "MECH1"
      ProcessValue <- "MantMS054"
   GraphicIOField "Campo ES gráfico_1" at 289,314 size 285x90; PictureList "BaseSullChico"
      ProcessValue <- "AnimaMS055"
   GraphicView "Visor de gráficos_2" at 333,200 size 201x179; Picture "secador_1"
   GraphicIOField "Campo ES gráfico_8" at 159,455 size 269x90; PictureList "BaseSullChico"
      ProcessValue <- "AnimaMS054"
   GraphicView "Visor de gráficos_4" at 333,200 size 201x179; Picture "Copia de secador"
      Visibility <- "MantMS055"
   GraphicView "Visor de gráficos_1" at 192,341 size 201x179; Picture "secador_1"
   GraphicView "Visor de gráficos_3" at 192,341 size 201x179; Picture "Copia de secador"
      Visibility <- "MantMS054"
   Button "Botón_3" at 1184,68 size 48x46; TextOff '?'
      on Click: ActivateScreen("MTA-AyudaSecBaja", 0)
   TextField "Campo de texto_1" at 527,9 size 226x27; Text 'Secadores de Baja presión'
   Button "Botón_18" at 639,277 size 200x82; TextOff 'Text'
      on Click: ActivateScreen("EPROC-BAJAMS055", 0)
   Button "Botón_1" at 482,410 size 200x82; TextOff 'Text'
      on Click: ActivateScreen("EPROC-BAJAMS054", 0)

screen "MTA-Sopladoras" 1280x800, template "Plantilla"
   Rectangle "Rectángulo_4" at 316,262 size 127x92
      Appearance <- "Sop1"
   IOField "Campo ES_1" at 301,378 size 151x31; Authorization "Administración de usuarios"; FormatPattern 9; Unit   Compresores
      ProcessValue <- "ReqSop1"
   IOField "Campo ES_2" at 492,378 size 153x31; Authorization "Administración de usuarios"; FormatPattern 9; Unit   Compresores
      ProcessValue <- "ReqSop2"
   IOField "Campo ES_3" at 691,378 size 153x31; Authorization "Administración de usuarios"; FormatPattern 9; Unit   Compresores
      ProcessValue <- "ReqSop3"
   IOField "Campo ES_4" at 766,443 size 90x23; FormatPattern 9
      ProcessValue <- "CompReqINI"
   TextField "Campo de texto_1" at 356,442 size 403x27; Text 'Cantidad de compresores que deben marchar:'
   TextField "Campo de texto_2" at 328,211 size 104x27; Text 'Sopladora 1'
   Button "Botón_12" at 1105,638 size 160x49; TextOff 'Volver'
      on Click: function_efd93a16()
   Button "Botón_1" at 323,269 size 112x38; TextOff 'Activar'; Authorization "Operación"
      on Click: SetBit("Sop1")
   Button "Botón_2" at 323,309 size 112x38; TextOff 'Desactivar'; Authorization "Operación"
      on Click: ResetBit("Sop1")
   Rectangle "Rectángulo_5" at 506,262 size 127x92
      Appearance <- "Sop2"
   Button "Botón_3" at 513,269 size 112x38; TextOff 'Activar'; Authorization "Operación"
      on Click: SetBit("Sop2")
   Button "Botón_4" at 513,309 size 112x38; TextOff 'Desactivar'; Authorization "Operación"
      on Click: ResetBit("Sop2")
   Rectangle "Rectángulo_6" at 704,262 size 127x92
      Appearance <- "Sop3"
   Button "Botón_5" at 711,269 size 112x38; TextOff 'Activar'; Authorization "Operación"
      on Click: SetBit("Sop3")
   Button "Botón_6" at 711,309 size 112x38; TextOff 'Desactivar'; Authorization "Operación"
      on Click: ResetBit("Sop3")
   TextField "Campo de texto_3" at 518,211 size 104x27; Text 'Sopladora 2'
   TextField "Campo de texto_4" at 716,211 size 104x27; Text 'Sopladora 3'
   TextField "Campo de texto_7" at 522,9 size 236x27; Text 'Seteo de sopladoras Activas'

